   TextField "Screen title" at 783,728 size 496x50; Text 'Screen title'
   Bar "Bar_1" at 262,206 size 122x241; MinimumValue 0; MaximumValue 100
      ProcessValue <- "20_TANKS_IP_DATA_RIO_06_FIRST_TANK_BWT_LEVEL"
   Button "Button_48" at 273,396 size 100x25; TextOff 'DISABLED'
      on Release: function_efd93a16("Tank 6P Status", 168, 315, -1, 2, 1)
      Visibility <- "504_Tank Grouping_DB2020_GROUP of TANK 12"
   Circle "Circle_3" at 340,212 size 14x14
      Appearance <- "20_TANKS_IP_DATA_RIO_06_FIRST_TANK_BWT_LEVEL_HIHI"
   TextField "Text field_125" at 295,212 size 51x14; Text 'LS425-6P'
   Polyline "Polyline_1" at 261,205 size 123x240
      Visibility <- "504_Tank Grouping_DB2020_RUN TANK 12"
   TextField "Text field_64" at 288,273 size 74x20; Text 'Tank - 6P'
   Bar "Bar_2" at 394,206 size 122x241; MinimumValue 0; MaximumValue 100
      ProcessValue <- "20_TANKS_IP_DATA_RIO_05_FIRST_TANK_BWT_LEVEL"
   Button "Button_44" at 406,396 size 100x25; TextOff 'DISABLED'
      on Release: function_efd93a16("Tank 5P Status", 168, 315, -1, 2, 1)
      Visibility <- "504_Tank Grouping_DB2020_GROUP of TANK 10"
   Circle "Circle_4" at 472,212 size 14x14
      Appearance <- "20_TANKS_IP_DATA_RIO_05_FIRST_TANK_BWT_LEVEL_HIHI"
   TextField "Text field_124" at 427,212 size 51x14; Text 'LS425-5P'
   Polyline "Polyline_2" at 392,205 size 123x240
      Visibility <- "504_Tank Grouping_DB2020_RUN TANK 10"
   TextField "Text field_8" at 418,275 size 74x20; Text 'Tank - 5P'
   Bar "Bar_3" at 525,206 size 122x241; MinimumValue 0; MaximumValue 100
      ProcessValue <- "20_TANKS_IP_DATA_RIO_04_FIRST_TANK_BWT_LEVEL"
   Button "Button_40" at 537,395 size 100x25; TextOff 'DISABLED'
      on Release: function_efd93a16("Tank 4P Status", 168, 315, -1, 2, 1)
      Visibility <- "504_Tank Grouping_DB2020_GROUP of TANK 8"
   Circle "Circle_5" at 604,212 size 14x14
      Appearance <- "20_TANKS_IP_DATA_RIO_04_FIRST_TANK_BWT_LEVEL_HIHI"
   TextField "Text field_123" at 559,212 size 51x14; Text 'LS425-4P'
   Polyline "Polyline_3" at 525,205 size 123x240
      Visibility <- "504_Tank Grouping_DB2020_RUN TANK 8"
   TextField "Text field_9" at 553,275 size 74x20; Text 'Tank - 4P'
   Bar "Bar_4" at 657,206 size 122x241; MinimumValue 0; MaximumValue 100
      ProcessValue <- "20_TANKS_IP_DATA_RIO_03_FIRST_TANK_BWT_LEVEL"
   Button "Button_36" at 668,395 size 100x25; TextOff 'DISABLED'
      on Release: function_efd93a16("Tank 3P Status", 168, 315, -1, 0, 1)
      Visibility <- "504_Tank Grouping_DB2020_GROUP of TANK 6"
   Circle "Circle_7" at 736,212 size 14x14
      Appearance <- "20_TANKS_IP_DATA_RIO_03_FIRST_TANK_BWT_LEVEL_HIHI"
   TextField "Text field_122" at 691,212 size 51x14; Text 'LS425-3P'
   Polyline "Polyline_4" at 656,205 size 123x240
      Visibility <- "504_Tank Grouping_DB2020_RUN TANK 6"
   TextField "Text field_14" at 680,275 size 74x20; Text 'Tank - 3P'
   Bar "Bar_5" at 789,206 size 122x241; MinimumValue 0; MaximumValue 100
      ProcessValue <- "20_TANKS_IP_DATA_RIO_02_FIRST_TANK_BWT_LEVEL"
   Button "Button_32" at 802,396 size 100x25; TextOff 'DISABLED'
      on Release: function_efd93a16("Tank 2P Status", 168, 315, -1, 0, 1)
      Visibility <- "504_Tank Grouping_DB2020_GROUP of TANK 4"
   Circle "Circle_15" at 868,212 size 14x14
      Appearance <- "20_TANKS_IP_DATA_RIO_02_FIRST_TANK_BWT_LEVEL_HIHI"
   TextField "Text field_121" at 823,212 size 51x14; Text 'LS425-2P'
   Polyline "Polyline_5" at 789,205 size 123x240
      Visibility <- "504_Tank Grouping_DB2020_RUN TANK 4"
   TextField "Text field_15" at 816,275 size 74x20; Text 'Tank - 2P'
   Bar "Bar_6" at 922,205 size 122x241; MinimumValue 0; MaximumValue 100
      ProcessValue <- "20_TANKS_IP_DATA_RIO_01_SECOND_TANK_BWT_LEVEL"
   Button "Button_52" at 934,395 size 100x25; TextOff 'DISABLED'
      on Release: function_efd93a16("Tank 1P Status", 168, 315, -1, 0, 1)
      Visibility <- "504_Tank Grouping_DB2020_GROUP of TANK 2"
   Circle "Circle_16" at 999,211 size 14x14
      Appearance <- "20_TANKS_IP_DATA_RIO_01_SECOND_TANK_BWT_LEVEL_HIHI"
   TextField "Text field_120" at 955,211 size 51x14; Text 'LS425-1P'
   Polyline "Polyline_6" at 921,205 size 123x240
      Visibility <- "504_Tank Grouping_DB2020_RUN TANK 2"
   GraphicView "Graphic view_6" at 127,446 size 591x12; Picture "Graphic_151"
   TextField "Text field_16" at 947,275 size 74x20; Text 'Tank - 1P'
   Bar "Bar_7" at 1096,334 size 122x241; MinimumValue 0; MaximumValue 100
      ProcessValue <- "20_TANKS_IP_DATA_RIO_01_FIRST_TANK_BWT_LEVEL"
   Circle "Circle_24" at 1168,339 size 14x14
      Appearance <- "20_TANKS_IP_DATA_RIO_01_FIRST_TANK_BWT_LEVEL_HIHI"
   TextField "Text field_133" at 1139,339 size 35x14; Text 'LS425'
   Polyline "Polyline_14" at 1095,332 size 125x242
      Visibility <- "504_Tank Grouping_DB2020_RUN TANK 1"
   Button "Button_56" at 1110,524 size 100x25; TextOff 'DISABLED'
      on Release: function_efd93a16("Tank FP Status", 168, 315, -1, 0, 1)
      Visibility <- "504_Tank Grouping_DB2020_GROUP of TANK 1"
   TextField "Text field_17" at 1111,400 size 111x20; Text 'Fore PeakTank'
   Bar "Bar_8" at 922,458 size 122x258; MinimumValue 0; MaximumValue 100
      ProcessValue <- "20_TANKS_IP_DATA_RIO_01_THIRD_TANK_BWT_LEVEL"
   Button "Button_54" at 933,661 size 100x25; TextOff 'DISABLED'
      on Release: function_efd93a16("Tank 1S Status", 168, 315, -1, 0, 1)
      Visibility <- "504_Tank Grouping_DB2020_GROUP of TANK 3"
   Circle "Circle_23" at 1000,464 size 14x14
      Appearance <- "20_TANKS_IP_DATA_RIO_01_THIRD_TANK_BWT_LEVEL_HIHI"
   TextField "Text field_126" at 955,465 size 51x14; Text 'LS422-1S'
   Polyline "Polyline_7" at 921,458 size 123x259
      Visibility <- "504_Tank Grouping_DB2020_RUN TANK 3"
   TextField "Text field_10" at 950,618 size 74x20; Text 'Tank - 1S'
   Bar "Bar_9" at 790,459 size 122x258; MinimumValue 0; MaximumValue 100
      ProcessValue <- "20_TANKS_IP_DATA_RIO_02_SECOND_TANK_BWT_LEVEL"
   Button "Button_34" at 801,662 size 100x25; TextOff 'DISABLED'
      on Release: function_efd93a16("Tank 2S Status", 168, 315, -1, 0, 1)
      Visibility <- "504_Tank Grouping_DB2020_GROUP of TANK 5"
   Circle "Circle_22" at 868,465 size 14x14
      Appearance <- "20_TANKS_IP_DATA_RIO_02_SECOND_TANK_BWT_LEVEL_HIHI"
   TextField "Text field_127" at 823,466 size 51x14; Text 'LS422-2S'
   Polyline "Polyline_8" at 789,458 size 123x259
      Visibility <- "504_Tank Grouping_DB2020_RUN TANK 5"
   TextField "Text field_11" at 817,618 size 74x20; Text 'Tank - 2S'
   Bar "Bar_10" at 659,460 size 122x258; MinimumValue 0; MaximumValue 100
      ProcessValue <- "20_TANKS_IP_DATA_RIO_03_SECOND_TANK_BWT_LEVEL"
   Button "Button_38" at 669,663 size 100x25; TextOff 'DISABLED'
      on Release: function_efd93a16("Tank 3S Status", 168, 315, -1, 0, 1)
      Visibility <- "504_Tank Grouping_DB2020_GROUP of TANK 7"
   Circle "Circle_21" at 736,467 size 14x14
      Appearance <- "20_TANKS_IP_DATA_RIO_03_SECOND_TANK_BWT_LEVEL_HIHI"
   TextField "Text field_128" at 691,468 size 51x14; Text 'LS422-3S'
   Polyline "Polyline_9" at 658,458 size 123x259
      Visibility <- "504_Tank Grouping_DB2020_RUN TANK 7"
   TextField "Text field_12" at 690,618 size 74x20; Text 'Tank - 3S'
   Bar "Bar_11" at 526,459 size 122x258; MinimumValue 0; MaximumValue 100
      ProcessValue <- "20_TANKS_IP_DATA_RIO_04_SECOND_TANK_BWT_LEVEL"
   Button "Button_42" at 537,662 size 100x25; TextOff 'DISABLED'
      on Release: function_efd93a16("Tank 4S Status", 168, 315, -1, 2, 1)
      Visibility <- "504_Tank Grouping_DB2020_GROUP of TANK 9"
   Circle "Circle_19" at 604,466 size 14x14
      Appearance <- "20_TANKS_IP_DATA_RIO_04_SECOND_TANK_BWT_LEVEL_HIHI"
   TextField "Text field_129" at 559,467 size 51x14; Text 'LS422-4S'
   Polyline "Polyline_10" at 525,458 size 123x259
      Visibility <- "504_Tank Grouping_DB2020_RUN TANK 9"
   TextField "Text field_13" at 554,618 size 74x20; Text 'Tank - 4S'
   Bar "Bar_12" at 394,459 size 122x258; MinimumValue 0; MaximumValue 100
      ProcessValue <- "20_TANKS_IP_DATA_RIO_05_SECOND_TANK_BWT_LEVEL"
   Button "Button_46" at 405,662 size 100x25; TextOff 'DISABLED'
      on Release: function_efd93a16("Tank 5S Status", 168, 315, -1, 2, 1)
      Visibility <- "504_Tank Grouping_DB2020_GROUP of TANK 11"
   Circle "Circle_18" at 472,465 size 14x14
      Appearance <- "20_TANKS_IP_DATA_RIO_05_SECOND_TANK_BWT_LEVEL_HIHI"
   TextField "Text field_130" at 427,466 size 51x14; Text 'LS422-5S'
   Polyline "Polyline_11" at 393,458 size 123x259
      Visibility <- "504_Tank Grouping_DB2020_RUN TANK 11"
   TextField "Text field_18" at 424,618 size 74x20; Text 'Tank - 5S'
   Bar "Bar_13" at 262,460 size 122x258; MinimumValue 0; MaximumValue 100
      ProcessValue <- "20_TANKS_IP_DATA_RIO_06_SECOND_TANK_BWT_LEVEL"
   Button "Button_50" at 273,663 size 100x25; TextOff 'DISABLED'
      on Release: function_efd93a16("Tank 6S Status", 168, 315, -1, 2, 1)
      Visibility <- "504_Tank Grouping_DB2020_GROUP of TANK 13"
   Circle "Circle_17" at 340,467 size 14x14
      Appearance <- "20_TANKS_IP_DATA_RIO_06_SECOND_TANK_BWT_LEVEL_HIHI"
   TextField "Text field_131" at 295,468 size 51x14; Text 'LS422-6S'
   Polyline "Polyline_12" at 261,458 size 123x258
      Visibility <- "504_Tank Grouping_DB2020_RUN TANK 13"
   TextField "Text field_19" at 290,618 size 74x20; Text 'Tank - 6S'
   Bar "Bar_14" at 39,324 size 119x258; Unit %; MinimumValue 0; MaximumValue 100
      ProcessValue <- "20_TANKS_IP_DATA_RIO_07_FIRST_TANK_BWT_LEVEL"
   Circle "Circle_25" at 108,330 size 14x14
      Appearance <- "20_TANKS_IP_DATA_RIO_07_FIRST_TANK_BWT_LEVEL_HIHI"
   TextField "Text field_132" at 79,330 size 35x14; Text 'LS425'
   Polyline "Polyline_13" at 38,324 size 121x259
      Visibility <- "504_Tank Grouping_DB2020_RUN TANK 14"
   Button "Button_58" at 48,527 size 100x25; TextOff 'DISABLED'
      on Release: function_efd93a16("Tank AP Status", 168, 315, -1, 2, 1)
      Visibility <- "504_Tank Grouping_DB2020_GROUP of TANK 14"
   Button "HmiScreenItemData_6" at 1043,144 size 116x50; TextOn 'Back'; TextOff 'Tank Status'
      on Release: ActivateScreen("Balast Water Treatment Plant", 0)
   Button "Button_2" at 252,437 size 37x30; TextOff 'DB&B'
      on Release: function_efd93a16("Double Block & Bleed Valve Monitoring", 250, 250, -1, -1, 1)
      Appearance <- "10_DI_DATA_CV407_OPN"
   TextField "Text field_65" at 190,398 size 46x25; Text 'PGC'
   TextField "Text field_75" at 183,480 size 60x20; Text 'Disabled'
   TextField "Text field_76" at 183,480 size 60x20; Text 'Enabled'
      Visibility <- "10_DI_DATA_E_400_RUN"
   GraphicView "Graphic view_76" at 185,421 size 57x55; Picture "Graphic_251"
   Button "Button_6" at 179,402 size 70x105; TextOff 'Text'
      on Release: ActivateScreen("PGC System", 0)
   TextField "Text field_20" at 53,396 size 103x20; Text 'Aft PeakTank'
   GraphicView "Graphic view_108" at 4,683 size 96x48; Picture "Left Arow"
   Button "HmiScreenItemData_14" at 3,660 size 106x93; TextOn 'Back'; TextOff 'Text'
      on Press: ActivateScreen("Inert Gas Conditioning Plant", 0)
   IOField "I/O field_1" at 68,460 size 84x25; FormatPattern 99.99; Unit m
      ProcessValue <- "Data_From_WBT_Level_APT m"
   IOField "I/O field_2" at 285,331 size 84x25; FormatPattern 99.99; Unit m
      ProcessValue <- "Data_From_WBT_Level_WBT_6P m"
   IOField "I/O field_3" at 418,331 size 84x25; FormatPattern 99.99; Unit m
      ProcessValue <- "Data_From_WBT_Level_WBT_5P m"
   IOField "I/O field_4" at 550,331 size 84x25; FormatPattern 99.99; Unit m
      ProcessValue <- "Data_From_WBT_Level_WBT_4P m"
   IOField "I/O field_5" at 681,331 size 84x25; FormatPattern 99.99; Unit m
      ProcessValue <- "Data_From_WBT_Level_WBT_3P m"
   IOField "I/O field_6" at 815,331 size 84x25; FormatPattern 99.99; Unit m
      ProcessValue <- "Data_From_WBT_Level_WBT_2P m"
   IOField "I/O field_7" at 949,331 size 84x25; FormatPattern 99.99; Unit m
      ProcessValue <- "Data_From_WBT_Level_WBT_1P m"
   IOField "I/O field_8" at 1124,459 size 84x25; FormatPattern 99.99; Unit m
      ProcessValue <- "Data_From_WBT_Level_FPT m"
   IOField "I/O field_9" at 945,555 size 84x25; FormatPattern 99.99; Unit m
      ProcessValue <- "Data_From_WBT_Level_WBT_1S m"
   IOField "I/O field_10" at 816,556 size 84x25; FormatPattern 99.99; Unit m
      ProcessValue <- "Data_From_WBT_Level_WBT_2S m"
   IOField "I/O field_11" at 685,558 size 84x25; FormatPattern 99.99; Unit m
      ProcessValue <- "Data_From_WBT_Level_WBT_3S m"
   IOField "I/O field_12" at 553,557 size 84x25; FormatPattern 99.99; Unit m
      ProcessValue <- "Data_From_WBT_Level_WBT_4S m"
   IOField "I/O field_13" at 418,558 size 84x25; FormatPattern 99.99; Unit m
      ProcessValue <- "Data_From_WBT_Level_WBT_5S m"
   IOField "I/O field_14" at 287,559 size 84x25; FormatPattern 99.99; Unit m
      ProcessValue <- "Data_From_WBT_Level_WBT_6S m"
   Button "Button_88" at 34,324 size 127x264; TextOff 'Text'
      on Release: function_efd93a16("Tank AP Status", 168, 315, -1, 0, 1)
      Appearance <- "504_Tank Grouping_DB2020_RUN TANK 14"
   Button "Button_86" at 259,458 size 126x260; TextOff 'Text'
      on Release: function_efd93a16("Tank 6S Status", 168, 315, -1, 0, 1)
      Appearance <- "504_Tank Grouping_DB2020_RUN TANK 13"
   Button "Button_79" at 391,457 size 126x262; TextOff 'Text'
      on Release: function_efd93a16("Tank 5S Status", 168, 315, -1, 0, 1)
      Appearance <- "504_Tank Grouping_DB2020_RUN TANK 11"
   Button "Button_77" at 523,457 size 126x262; TextOff 'Text'
      on Release: function_efd93a16("Tank 4S Status", 168, 315, -1, 0, 1)
      Appearance <- "504_Tank Grouping_DB2020_RUN TANK 9"
   Button "Button_74" at 657,457 size 126x262; TextOff 'Text'
      on Release: function_efd93a16("Tank 3S Status", 168, 315, -1, 0, 1)
      Appearance <- "504_Tank Grouping_DB2020_RUN TANK 7"
   Button "Button_70" at 788,457 size 126x262; TextOff 'Text'
      on Release: function_efd93a16("Tank 2S Status", 168, 315, -1, 0, 1)
      Appearance <- "504_Tank Grouping_DB2020_RUN TANK 5"
   Button "Button_66" at 921,457 size 126x261; TextOff 'Text'
      on Release: function_efd93a16("Tank 1S Status", 168, 315, -1, 0, 1)
      Appearance <- "504_Tank Grouping_DB2020_RUN TANK 3"
   Button "Button_61" at 1093,328 size 130x248; TextOff 'Text'
      on Release: function_efd93a16("Tank FP Status", 168, 315, -1, 0, 1)
      Appearance <- "504_Tank Grouping_DB2020_RUN TANK 1"
   Button "Button_62" at 919,205 size 126x242; TextOff 'Text'
      on Release: function_efd93a16("Tank 1P Status", 168, 315, -1, 0, 1)
      Appearance <- "504_Tank Grouping_DB2020_RUN TANK 2"
   Button "Button_68" at 789,202 size 126x246; TextOff 'Text'
      on Release: function_efd93a16("Tank 2P Status", 168, 315, -1, 0, 1)
      Appearance <- "504_Tank Grouping_DB2020_RUN TANK 4"
   Button "Button_72" at 654,205 size 126x242; TextOff 'Text'
      on Release: function_efd93a16("Tank 3P Status", 168, 315, -1, 0, 1)
      Appearance <- "504_Tank Grouping_DB2020_RUN TANK 6"
   Button "Button_76" at 524,205 size 126x243; TextOff 'Text'
      on Release: function_efd93a16("Tank 4P Status", 168, 315, -1, 0, 1)
      Appearance <- "504_Tank Grouping_DB2020_RUN TANK 8"
   Button "Button_78" at 392,206 size 126x241; TextOff 'Text'
      on Release: function_efd93a16("Tank 5P Status", 168, 315, -1, 0, 1)
      Appearance <- "504_Tank Grouping_DB2020_RUN TANK 10"
   Button "Button_84" at 259,204 size 126x244; TextOff 'Text'
      on Release: function_efd93a16("Tank 6P Status", 168, 315, -1, 0, 1)
      Appearance <- "504_Tank Grouping_DB2020_RUN TANK 12"
   Group "Group_5" at 664,46 size 45x27; FormatPattern 999
   Group "Group_1" at 711,46 size 50x27; FormatPattern 999; Unit h
   Group "Group_2" at 605,46 size 57x27; FormatPattern 999; Unit h
   Button "HmiScreenItemData_5" at 180,144 size 116x50; TextOn 'Back'; TextOff 'Tank Status'
      on Release: function_efd93a16("Tank Status", 400, 250, -1, -1, 1)
   Button "Button_10" at 14,93 size 153x55; TextOff 'Text'
      on Release: function_efd93a16("Salinity - Acceptance", 168, 315, -1, 0, 1)
      Visibility <- "2068_Sys_Status_Data_SAL_VALID"
   Button "Button_12" at 14,93 size 153x53; TextOff 'Text'
      on Release: function_efd93a16("Tank Times", 300, 200, -1, 0, 1)
      Visibility <- "2068_Sys_Status_Data_Times Visibil"
   Button "Button_59" at 298,44 size 240x30; TextOn 'TB3 Enabled'; TextOff 'BWT System Shutting Down'
      Visibility <- "2110_BTCS_CNTRL_DB_BTCS_STATE"
   Button "Button_60" at 299,44 size 240x30; TextOn 'TB3 Enabled'; TextOff 'BWT System Enabled'
      Visibility <- "2110_BTCS_CNTRL_DB_BTCS_STATE"
   IOField "I/O field_29" at 664,46 size 45x27; FormatPattern 99; Unit h
      ProcessValue <- "Sequence Times_DB_Treatment Timer_Hours Left"
      Visibility <- "2110_BTCS_CNTRL_DB_BTCS_STATE"
   IOField "I/O field_30" at 664,46 size 45x27; FormatPattern 99; Unit h
      ProcessValue <- "Sequence Times_DB_Pre-Dwell Timer_Hours Left"
      Visibility <- "2110_BTCS_CNTRL_DB_BTCS_STATE"
   IOField "I/O field_15" at 711,46 size 50x27; FormatPattern 99; Unit m
      ProcessValue <- "Sequence Times_DB_Treatment Timer_Minutes Left"
      Visibility <- "2110_BTCS_CNTRL_DB_BTCS_STATE"
   IOField "I/O field_16" at 711,46 size 50x27; FormatPattern 99; Unit m
      ProcessValue <- "Sequence Times_DB_Pre-Dwell Timer_Minutes Left"
      Visibility <- "2110_BTCS_CNTRL_DB_BTCS_STATE"
   IOField "I/O field_17" at 605,46 size 57x27; FormatPattern 999; Unit d
      ProcessValue <- "Sequence Times_DB_Treatment Timer_Days Left"
      Visibility <- "2110_BTCS_CNTRL_DB_BTCS_STATE"
   IOField "I/O field_18" at 605,46 size 57x27; FormatPattern 999; Unit d
      ProcessValue <- "Sequence Times_DB_Pre-Dwell Timer_Days Left"
      Visibility <- "2110_BTCS_CNTRL_DB_BTCS_STATE"

screen "PGC System" 1280x800, template "Template"
   Button "HmiScreenItemData_1" at -189,1 size 150x43; TextOn 'Back'; TextOff 'Main Index'
      on Release: ActivateScreen("02 Main Index", 0)
   Gauge "Gauge_1" at 454,351 size 184x184; CaptionText 'Pressure'; UnitText 'Bar'
      ProcessValue <- "12_AI_Data_E_400_PT002_SCALED"
      MaximumValue <- "84_Setpoints_E400_PT002_HighHigh"
   TextField "Text field_20" at 187,312 size 324x26; Text 'Process Gas Discharge Pressure'
   TextField "Text field_7" at 221,72 size 326x26; Text 'Process Gas Compressor Control'
   TextField "Text field_10" at 119,405 size 243x20; Text 'Process Gas Discharge Pressure'
   TextField "Text field_17" at 119,464 size 217x20; Text 'Discharge Pressure Setpoint'
   Button "Button_8" at 117,115 size 240x30; TextOn 'TB3 Enabled'; TextOff 'PGC System Not Running OK'
      Visibility <- "10_DI_DATA_E_400_RUN"
   Button "HmiScreenItemData_12" at 141,237 size 69x51; TextOn 'Back'; TextOff 'Reset'; Authorization "Operate"
      on Press: function_b14e0dd5("140_PGC_HRS_RUN_DB_RST", 0)
   IOField "I/O field_10" at 70,236 size 66x25; FormatPattern 9999; Unit  h
      ProcessValue <- "140_PGC_HRS_RUN_DB_SRV_HRS"
   TextField "Text field_22" at 36,238 size 37x20; Text 'Run'
   TextField "Text field_23" at 36,268 size 37x20; Text 'Set'
   TextField "Text field_24" at 79,212 size 100x20; Text 'Service Hour'
   IOField "I/O field_13" at 222,249 size 75x25; FormatPattern 99999; Unit h
      ProcessValue <- "140_PGC_HRS_RUN_DB_HRS"
   IOField "I/O field_14" at 299,249 size 40x25; FormatPattern 99; Unit m
      ProcessValue <- "140_PGC_HRS_RUN_DB_MINS"
   IOField "I/O field_15" at 341,249 size 40x25; FormatPattern 99; Unit s
      ProcessValue <- "140_PGC_HRS_RUN_DB_SECS"
   Button "Button_7" at 654,76 size 57x25; TextOn 'Alarm'; TextOff 'Service'
      Visibility <- "140_PGC_HRS_RUN_DB_SRVC"
      Appearance <- "140_PGC_HRS_RUN_DB_SRVC"
   Button "Button_15" at 187,173 size 57x25; TextOn 'Enabled'; TextOff 'Disabled'
   Button "Button_16" at 341,173 size 64x25; TextOn 'Alarm'; TextOff 'Text'
   TextField "Text field_14" at 44,175 size 115x20; Text 'PG Compressor'
   TextField "Text field_15" at 191,151 size 60x18; Text 'Enabled'
   TextField "Text field_16" at 266,151 size 64x18; Text 'Running'
   TextField "Text field_18" at 343,150 size 78x18; Text 'Shutdown'
   Button "Button_1" at 264,173 size 57x25; TextOn 'Enabled'; TextOff 'Stopped'
   TextField "Text field_32" at 187,173 size 57x25; Text 'Enabled'
      Visibility <- "10_DI_DATA_E_400_SHTDN"
   TextField "Text field_2" at 264,173 size 57x25; Text 'Running'
      Visibility <- "10_DI_DATA_E_400_RUN"
   Button "Button_3" at 341,173 size 64x25; TextOn 'Enabled'; TextOff 'Normal'
   Button "Button_2" at 341,173 size 69x25; TextOn 'Alarm'; TextOff 'Shutdown'
      Visibility <- "10_DI_DATA_E_400_NOK"
      Appearance <- "10_DI_DATA_E_400_NOK"
   Gauge "Gauge_2" at 454,588 size 184x184; UnitText '°C'; CaptionText 'Temperature'
      ProcessValue <- "12_AI_Data_E_400_TE002_SCALED"
      MaximumValue <- "84_Setpoints_E400_TT002_HighHigh"
   TextField "Text field_1" at 187,549 size 365x26; Text 'Process Gas Discharge Temperature'
   TextField "Text field_3" at 119,641 size 178x20; Text 'Discharge Temperature'
   TextField "Text field_4" at 109,699 size 246x20; Text 'Discharge Temperature Setpoint'
   IOField "I/O field_2" at 332,403 size 66x25; FormatPattern 9.99; Unit  Bar
      ProcessValue <- "12_AI_Data_E_400_PT002_SCALED"
   IOField "I/O field_1" at 334,638 size 66x25; FormatPattern 999; Unit  °C
      ProcessValue <- "12_AI_Data_E_400_TE002_SCALED"
   Button "HmiScreenItemData_11" at 3,1 size 150x43; TextOn 'IGG Plant'; TextOff 'GCU Plant'
      on Release: ActivateScreen("Inert Gas Conditioning Plant", 0)
   IOField "I/O field_3" at 332,462 size 66x25; Authorization "Commissioning"; FormatPattern 9.99; Unit  Bar
      ProcessValue <- "84_Setpoints_E400_PT002_HighHigh"
   IOField "I/O field_4" at 334,697 size 66x25; Authorization "Commissioning"; FormatPattern 999; Unit  °C
      ProcessValue <- "84_Setpoints_E400_TT002_HighHigh"
   GraphicView "Graphic view_1" at 514,109 size 192x199; Picture "Graphic_251"
   Button "HmiScreenItemData_3" at 1125,1 size 150x43; TextOn 'I&A Compressor Ok'; TextOff 'Back'
      on Release: function_efd93a16()
   TextField "Text field_5" at 222,226 size 160x25; Text 'Total Run Time'
   TextField "Text field_6" at 818,74 size 312x26; Text 'Process Gas Compressor Purge'
   TextField "Text field_8" at 717,177 size 263x20; Text 'Process Gas Compresor Stop Delay'
   TextField "Text field_11" at 716,111 size 305x20; Text 'Combustion Air Blower after Start Delay'
   IOField "I/O field_7" at 993,109 size 66x25; FormatPattern 999; Unit s
      ProcessValue <- "PGC Flush_DB_CAB after Start Delay"
   TextField "Text field_12" at 716,144 size 208x20; Text 'Combustion Air Blower RPM'
   IOField "I/O field_8" at 993,142 size 66x25; FormatPattern 999; Unit RPM
      ProcessValue <- "PGC Flush_DB_CAB RPM Cmnd"
   Button "HmiScreenItemData_2" at 982,285 size 82x35; TextOn 'Back'; TextOff 'Override'; Authorization "Operating Mode"
      on Press: function_b14e0dd5("PGC Flush_DB_Override", 0)
      Appearance <- "PGC Flush_DB_Flip Flop_Override_Output"
   TextField "Text field_9" at 1068,149 size 91x21; Text 'Running'
      Appearance <- "PGC Flush_DB_Running"
   TextField "Text field_13" at 1068,129 size 91x21; Text 'Enabled'
      Appearance <- "PGC Flush_DB_Activate"
   TextField "Text field_19" at 1068,329 size 91x21; Text 'Done'
      Appearance <- "PGC Flush_DB_Done"
   TextField "Text field_21" at 1068,169 size 91x21; Text 'Open CV405'
      Appearance <- "PGC Flush_DB_CV405 Open"
   TextField "Text field_25" at 1068,189 size 91x21; Text 'Open CV401'
      Appearance <- "PGC Flush_DB_CV401 Open"
   TextField "Text field_26" at 1068,209 size 91x21; Text 'Open CV431'
      Appearance <- "PGC Flush_DB_CV431 Open"
   TextField "Text field_27" at 1068,249 size 91x21; Text 'Close CV441'
      Appearance <- "PGC Flush_DB_CV431 Open"
   TextField "Text field_28" at 1068,269 size 91x21; Text 'Start CAB'
      Appearance <- "PGC Flush_DB_CAB Start"
   TextField "Text field_29" at 1068,289 size 91x21; Text 'Mdlt CV403'
      Appearance <- "PGC Flush_DB_CV403 Modulate"
   TextField "Text field_30" at 1068,309 size 91x21; Text 'Stop PGC'
      Appearance <- "PGC Flush_DB_Stop PGC"
   IOField "I/O field_37" at 890,604 size 90x29; Authorization "Commissioning"; FormatPattern 999; Unit  step
      ProcessValue <- "2110_BTCS_CNTRL_DB_BTCS_STEP"
   Button "HmiScreenItemData_10" at 749,604 size 137x29; TextOn 'Back'; TextOff 'BWTS Step'
   Button "HmiScreenItemData_51" at 749,671 size 137x29; TextOn 'Back'; TextOff 'BWTS State'
   Button "HmiScreenItemData_54" at 749,633 size 495x29; TextOn 'Back'; TextOff 'IGG STEP'; TextList "STEP LIST BTCS"
      ProcessValue <- "2110_BTCS_CNTRL_DB_BTCS_STEP"
   Button "HmiScreenItemData_55" at 749,700 size 495x29; TextOn 'Back'; TextOff 'IGG STEP'; TextList "STATE LIST BTCS"
      ProcessValue <- "2110_BTCS_CNTRL_DB_BTCS_STATE"
   IOField "I/O field_38" at 890,671 size 90x29; Authorization "Commissioning"; FormatPattern 9; Unit  state
      ProcessValue <- "2110_BTCS_CNTRL_DB_BTCS_STATE"
   TextField "Text field_31" at 716,210 size 149x20; Text 'PGC Purge Duration'
   IOField "I/O field_6" at 993,208 size 66x25; FormatPattern 999; Unit m
      ProcessValue <- "PGC Flush_DB_PGC Purge Duration"
   TextField "Text field_33" at 1068,229 size 91x21; Text 'Open CV403'
      Appearance <- "PGC Flush_DB_CV403 Open"
   TextField "Text field_34" at 768,296 size 175x18; Text 'Purge Request Simulate'
      Visibility <- "user_group"
   Switch "Switch_1" at 726,288 size 32x29; CaptionText 'Switch'; TextOn 'ON'; TextOff 'OFF'; Authorization "User administration"; PictureOff "Design_5_PilotLight_Green_Off"; PictureOn "Design_5_PilotLight_Green_On"
      on Change: InvertBit("Sequence Times_DB_Treatment Timer_Enable")
      Visibility <- "user_group"
      ProcessValue <- "19_AUTO_CMNDS_Data_Purge Rqst Simulate"
   TextField "Text field_35" at 1160,149 size 106x21; Text 'Running'
      Appearance <- "PGC Flush_DB_Running"
   TextField "Text field_36" at 1160,129 size 106x21; Text 'Enabled'
      Appearance <- "PGC Flush_DB_Activate"
   TextField "Text field_37" at 1160,329 size 106x21; Text 'Done'
      Appearance <- "100_GCU_AUTO_SEQ_DB_CRNT_STEP"
   TextField "Text field_38" at 1160,169 size 106x21; Text 'Opened CV405'
      Appearance <- "1405_PID_CV405_ManualEnable"
   TextField "Text field_39" at 1160,189 size 106x21; Text 'Opened CV401'
      Appearance <- "PGC Flush_DB_CV401 Opened"
   TextField "Text field_40" at 1160,209 size 106x21; Text 'Opened CV431'
      Appearance <- "PGC Flush_DB_CV431 Opened"
   TextField "Text field_41" at 1160,249 size 106x21; Text 'Closed CV441'
      Appearance <- "PGC Flush_DB_CV441 Closed"
   TextField "Text field_42" at 1160,269 size 106x21; Text 'Started CAB'
      Appearance <- "PGC Flush_DB_CAB Started"
   TextField "Text field_43" at 1160,289 size 106x21; Text 'Mdling CV403'
      Appearance <- "1403_PID_300CV403_ModeActivate"
   TextField "Text field_44" at 1160,309 size 106x21; Text 'Stoped PGC'
      Appearance <- "PGC Flush_DB_PGC Stoped"
   TextField "Text field_45" at 1160,229 size 106x21; Text 'Opened CV403'
      Appearance <- "1403_PID_300CV403_ManualEnable"
   TextField "Text field_46" at 711,332 size 173x20; Text 'Air / Inert Gas Pressure'
   Button "Button_9" at 1001,329 size 57x25; TextOn 'Enabled'; TextOff 'Text'
   TextField "Text field_47" at 710,366 size 277x20; Text 'Air / Inert Gas Pressure Setpoint (Pre-Ignition)'
   Button "Button_11" at 1001,364 size 57x25; TextOn 'Enabled'; TextOff 'Text'
   TextField "Text field_48" at 718,498 size 182x20; Text 'Modulating Valve Position'
   TextField "Text field_49" at 709,399 size 278x20; Text 'Air / Inert Gas Pressure Setpoint (Main-Ignition)'
   Button "Button_10" at 1001,397 size 57x25; TextOn 'Enabled'; TextOff 'Text'
   IOField "I/O field_9" at 993,329 size 66x25; FormatPattern 999; Unit  mbar
      ProcessValue <- "12_AI_Data_PIT402_SCALED"
   IOField "I/O field_12" at 993,364 size 66x25; Authorization "Commissioning"; FormatPattern 999; Unit  mbar
      ProcessValue <- "84_Setpoints_PIT402_Pilot_Target"
   IOField "I/O field_16" at 993,495 size 66x25; FormatPattern 999; Unit  %
      ProcessValue <- "16_AQ_Data_CV403_CNTRL"
   IOField "I/O field_17" at 993,462 size 66x25; FormatPattern 999; Unit  mBar
      ProcessValue <- "19_AUTO_CMNDS_Data_PIT402_Target"
      Appearance <- "19_AUTO_CMNDS_Data_PIT402_Target"
   IOField "I/O field_18" at 993,396 size 66x25; Authorization "Commissioning"; FormatPattern 999; Unit  mbar
      ProcessValue <- "84_Setpoints_PIT402_Main_Target"
   TextField "Text field_50" at 1068,497 size 58x20; Text 'Opened'
   TextField "Text field_51" at 711,465 size 266x20; Text 'Air / Inert Gas Pressure Setpoint (Current)'
   TextField "Text field_52" at 709,432 size 278x20; Text 'Air / Inert Gas Pressure Setpoint (Post-Ignition)'
   Button "Button_4" at 1001,430 size 57x25; TextOn 'Enabled'; TextOff 'Text'
   IOField "I/O field_19" at 993,429 size 66x25; Authorization "Commissioning"; FormatPattern 999; Unit  mbar
      ProcessValue <- "84_Setpoints_PIT401_Post_Target_Max"
   TextField "Text field_53" at 1079,107 size 73x20; Text 'Command'
   TextField "Text field_54" at 1182,107 size 73x20; Text 'Feedback'
   IOField "I/O field_20" at 70,266 size 66x25; Authorization "Commissioning"; FormatPattern 9999; Unit h
      ProcessValue <- "140_PGC_HRS_RUN_DB_SHRS_IP"
   TextField "Text field_55" at 716,243 size 168x20; Text 'Temperature Setpoint'
   IOField "I/O field_11" at 993,241 size 66x25; FormatPattern 999; Unit  °C
      ProcessValue <- "PGC Flush_DB_Temperature Setpoint"
   Button "HmiScreenItemData_19" at 749,567 size 495x29; TextOn 'Back'; TextOff 'IGG STEP'; TextList "STEP LIST_GCU"
      ProcessValue <- "100_GCU_AUTO_SEQ_DB_CRNT_STEP"
   IOField "I/O field_21" at 890,537 size 90x29; Authorization "Commissioning"; FormatPattern 999; Unit  Step
      ProcessValue <- "100_GCU_AUTO_SEQ_DB_CRNT_STEP"
   Button "HmiScreenItemData_9" at 749,536 size 100x30; TextOn 'Back'; TextOff 'GCU PLC'
   Button "HmiScreenItemData_16" at 238,742 size 83x29; TextOn 'Back'; TextOff 'Temp-Trends'
      on Click: function_efd93a16("PGC Temperature Trends", 200, 100, -1, -1, 1)
   IOField "I/O field_22" at 993,175 size 66x25; FormatPattern 999; Unit m
      ProcessValue <- "PGC Flush_DB_PGC Stop Delay"

screen "Fresh Water System" 1280x800, template "Template"
   GraphicView "Graphic view_29" at 858,564 size 26x29; Picture "Graphic_155"
   Bar "Bar_1" at 145,436 size 311x274; Unit  %; MinimumValue 0; MaximumValue 100
      ProcessValue <- "12_AI_Data_LIT305_SCALED"
   GraphicView "Graphic view_15" at 640,691 size 216x15; Picture "Graphic_156"
   GraphicView "Graphic view_22" at 468,691 size 71x15; Picture "Graphic_156"
   TextField "Text field_1" at 262,720 size 73x32; Text 'IBC-2 Bulk Tank'
   GraphicView "Graphic view_3" at 454,688 size 6x20; Picture "Graphic_113"
   TextField "Text field_4" at 442,89 size 268x26; Text 'Fresh Water Pump Control'
   IOField "I/O field_2" at 646,242 size 65x25; FormatPattern 99999; Unit  h
      ProcessValue <- "P305_Functioning Hours_IDB_Hours Functioning Out"
   TextField "Text field_5" at 616,244 size 37x20; Text 'Run'
   TextField "Text field_6" at 616,275 size 37x20; Text 'Set'
   TextField "Text field_9" at 659,141 size 100x20; Text 'Service Hour'
   Button "HmiScreenItemData_10" at 639,169 size 178x34; TextOn 'Back'; TextOff 'Text'
   IOField "I/O field_4" at 689,173 size 40x25; FormatPattern 99; Unit h
      ProcessValue <- "82_To_HMI_P305 FW Pump Run Hours"
   IOField "I/O field_5" at 730,173 size 40x25; FormatPattern 99; Unit m
      ProcessValue <- "P305_Functioning Hours_IDB_Minutes"
   IOField "I/O field_6" at 771,173 size 40x25; FormatPattern 99; Unit s
      ProcessValue <- "P305_Functioning Hours_IDB_Seconds"
   Button "Button_4" at 776,90 size 57x25; TextOn 'Alarm'; TextOff 'Service'
      Visibility <- "P305_Functioning Hours_IDB_Service Time bit"
   Button "Button_9" at 374,166 size 57x25; TextOn 'Enabled'; TextOff 'Disabled'
   Button "Button_11" at 528,166 size 64x25; TextOn 'Alarm'; TextOff 'Text'
   TextField "Text field_10" at 231,168 size 140x20; Text 'Fresh Water Pump'
   TextField "Text field_8" at 378,144 size 60x18; Text 'Enabled'
   TextField "Text field_17" at 453,144 size 64x18; Text 'Running'
   TextField "Text field_20" at 533,144 size 58x18; Text 'Tripped'
      Visibility <- "10 DI_DATA_P305_TRIPPED(1)"
   Button "Button_12" at 451,166 size 57x25; TextOn 'Enabled'; TextOff 'Stopped'
   TextField "Text field_26" at 374,166 size 57x25; Text 'Enabled'
      Visibility <- "14_DQ_Data_P305ControlOut"
   TextField "Text field_27" at 448,166 size 64x25; Text 'Running'
      Visibility <- "10 DI_DATA_P305_ENBLD"
   GraphicView "Graphic view_12" at 396,411 size 20x26; Picture "Graphic_36"
   TextField "Text field_11" at 421,411 size 60x18; Text 'LIT-305'
   GraphicView "Graphic view_13" at 518,691 size 71x15; Picture "Graphic_156"
   GraphicView "Graphic view_11" at 456,691 size 15x15; Picture "Graphic_156"
   GraphicView "Graphic view_27" at 846,676 size 25x29; Picture "Graphic_153"
   GraphicView "Graphic view_28" at 858,581 size 13x101; Picture "Graphic_152"
   GraphicView "Graphic view_30" at 876,702 size 146x15; Picture "Graphic_156"
   GraphicView "Graphic view_31" at 870,564 size 152x15; Picture "Graphic_156"
   GraphicView "Graphic view_32" at 858,688 size 26x29; Picture "Graphic_166"
   TextField "Text field_15" at 550,746 size 133x32; Text 'P-305 Fresh Water Pump'
   Button "Button_1" at 528,166 size 64x25; TextOn 'Alarm'; TextOff 'Tripped'
      Visibility <- "10 DI_DATA_P305_TRIPPED"
      Appearance <- "10 DI_DATA_P305_TRIPPED"
   IOField "I/O field_13" at 376,388 size 63x18; FormatPattern 99.9; Unit  %
      ProcessValue <- "12_AI_Data_LIT305_SCALED"
   TextField "Text field_22" at 1059,560 size 168x21; Text 'Fresh Water Supply To GCU'
   TextField "Text field_3" at 1059,699 size 168x21; Text 'Fresh Water Supply To IGG'
   Button "HmiScreenItemData_9" at 721,243 size 69x51; TextOn 'Back'; TextOff 'SReset'; Authorization "Operating Mode"
      on Press: function_b14e0dd5("82_To_HMI_P305 FW Pump Reset Hours", 0)
   GraphicView "Graphic view_1" at 1021,697 size 32x24; Picture "Graphic_244"
   GraphicView "Graphic view_2" at 1021,558 size 32x24; Picture "Graphic_244"
   Button "HmiScreenItemData_1" at 1,1 size 150x43; TextOn 'Back'; TextOff 'Main Index'
      on Release: ActivateScreen("02 Main Index", 0)
   GraphicIOField "Graphic I/O field_3" at 586,670 size 60x65; PictureList "Pump Ani"
      ProcessValue <- "FW Pump Animation"
   Button "HmiScreenItemData_3" at 1129,1 size 150x43; TextOn 'I&A Compressor Ok'; TextOff 'Back'
      on Release: function_efd93a16()
   AlarmView "Alarm view_1" at 0,777 size 1280x23
   IOField "I/O field_21" at 617,211 size 90x25; FormatPattern 999999; Unit  h
      ProcessValue <- "P305_Functioning Hours_IDB_Hours Total"
      Visibility <- "80_From_HMI_P301_PRSNT"
   TextField "Text field_31" at 712,213 size 123x20; Text 'Total Run Hours'
      Visibility <- "80_From_HMI_P301_PRSNT"
   IOField "I/O field_1" at 648,173 size 40x25; FormatPattern 99; Unit d
      ProcessValue <- "82_To_HMI_P305 FW Pump Run Days"
   IOField "I/O field_9" at 646,273 size 65x25; Authorization "Commissioning"; FormatPattern 99999; Unit  h
      ProcessValue <- "82_To_HMI_P305 FW Pump Service Time Hours"
   Button "HmiScreenItemData_4" at 488,210 size 75x34; TextOn 'STOP'; TextOff 'Stop'
      on Press: ResetBit("80_From_HMI_MAN_DQ_1_7(1)")
   Button "HmiScreenItemData_2" at 385,210 size 75x34; TextOn 'START'; TextOff 'Start'
      on Press: SetBit("80_From_HMI_MAN_DQ_1_7(1)")
   Rectangle "Rectangle_7" at 208,78 size 656x250
      Visibility <- "80_From_HMI_P305_PRSNT"

screen "GCU Process Times" 1280x800, template "Template"
   on GenerateScreen: "TitleUpdater"()
   Button "HmiScreenItemData_1" at 1,1 size 150x43; TextOn 'Back'; TextOff 'Commissioning'
      on Release: ActivateScreen("Commissioning Main Page", 0)
   AlarmView "Alarm view_1" at 0,777 size 1280x23
   TextField "Text field_29" at 545,103 size 65x20; Text 'Time (s)'
   TextField "Text field_65" at 240,128 size 300x25; Text 'P303 Started Delay'
   TextField "Text field_42" at 240,103 size 89x20; Text 'Description'
   IOField "I/O field_128" at 545,128 size 65x25; Authorization "Parameter Change"; FormatPattern 999
      ProcessValue <- "86_Times_P303_STRTD_DLY"
   TextField "Text field_53" at 240,74 size 193x26; Text 'GCU Process Times'
   TextField "Text field_1" at 240,158 size 300x25; Text 'P303 Stopped Delay'
   IOField "I/O field_1" at 545,158 size 65x25; Authorization "Parameter Change"; FormatPattern 999
      ProcessValue <- "86_Times_P303_STPD_DLY"
   TextField "Text field_2" at 240,188 size 300x25; Text 'P304 Started Delay'
   IOField "I/O field_2" at 545,188 size 65x25; Authorization "Parameter Change"; FormatPattern 999
      ProcessValue <- "86_Times_P304_STRTD_DLY"
   TextField "Text field_3" at 240,218 size 300x25; Text 'P304 Stopped Delay'
   IOField "I/O field_3" at 545,218 size 65x25; Authorization "Parameter Change"; FormatPattern 999
      ProcessValue <- "86_Times_P304_STPD_DLY"
   TextField "Text field_4" at 240,248 size 300x25; Text 'P305 Started Delay'
   IOField "I/O field_4" at 545,248 size 65x25; Authorization "Parameter Change"; FormatPattern 999
      ProcessValue <- "86_Times_P305_STRTD_DLY"
   TextField "Text field_5" at 240,278 size 300x25; Text 'P305 Stopped Delay'
   IOField "I/O field_5" at 545,278 size 65x25; Authorization "Parameter Change"; FormatPattern 999
      ProcessValue <- "86_Times_P305_STPD_DLY"
   TextField "Text field_6" at 240,308 size 300x25; Text 'CV341 Closed Delay'
   IOField "I/O field_6" at 545,308 size 65x25; Authorization "Parameter Change"; FormatPattern 999
      ProcessValue <- "86_Times_CV341_CLSD_DLY"
   TextField "Text field_7" at 240,338 size 300x25; Text 'CV358 Closed Delay'
   IOField "I/O field_7" at 545,338 size 65x25; Authorization "Parameter Change"; FormatPattern 999
      ProcessValue <- "86_Times_CV358_CLSD_DLY"
   TextField "Text field_8" at 975,103 size 65x20; Text 'Time (s)'
   TextField "Text field_9" at 670,128 size 300x25; Text 'CV405 Opened Delay'
   TextField "Text field_10" at 670,103 size 89x20; Text 'Description'
   IOField "I/O field_8" at 975,128 size 65x25; Authorization "Parameter Change"; FormatPattern 999
      ProcessValue <- "86_Times_CV405_OPND_DLY"
   TextField "Text field_11" at 670,158 size 300x25; Text 'CV406 Closed Delay'
   IOField "I/O field_9" at 975,158 size 65x25; Authorization "Parameter Change"; FormatPattern 999
      ProcessValue <- "86_Times_CV406_CLSD_DLY"
   TextField "Text field_12" at 670,188 size 300x25; Text 'E400 Stop Time'
   IOField "I/O field_10" at 975,188 size 65x25; Authorization "Parameter Change"; FormatPattern 999
      ProcessValue <- "86_Times_E400_STOP_TIME"
   TextField "Text field_13" at 670,218 size 300x25; Text 'P303 Stop Time'
   IOField "I/O field_11" at 975,218 size 65x25; Authorization "Parameter Change"; FormatPattern 999
      ProcessValue <- "86_Times_P303_STOP_TIME"
   TextField "Text field_14" at 670,248 size 300x25; Text 'CV341 Opened Delay'
   IOField "I/O field_12" at 975,248 size 65x25; Authorization "Parameter Change"; FormatPattern 999
      ProcessValue <- "86_Times_CV341_OPND_DLY"
   TextField "Text field_15" at 670,278 size 300x25; Text 'GCU Tank Maximum Drain Time'
   IOField "I/O field_13" at 975,278 size 65x25; Authorization "Parameter Change"; FormatPattern 999
      ProcessValue <- "86_Times_GCU_TNK_DRN_MAX_TIME"
   TextField "Text field_16" at 670,308 size 300x25; Text 'GCU Flush Time'
   IOField "I/O field_14" at 975,308 size 65x25; Authorization "Parameter Change"; FormatPattern 999
      ProcessValue <- "86_Times_GCU_FLUSH_TIME"
   TextField "Text field_17" at 670,338 size 300x25; Text 'Post Flush Delay'
   IOField "I/O field_15" at 975,338 size 65x25; Authorization "Parameter Change"; FormatPattern 999
      ProcessValue <- "86_Times_POST_FLUSH_DLY"
   TextField "Text field_18" at 240,368 size 300x25; Text 'CV401 Opened Delay'
   IOField "I/O field_16" at 545,368 size 65x25; Authorization "Parameter Change"; FormatPattern 999
      ProcessValue <- "86_Times_CV401_OPND_DLY"
   TextField "Text field_19" at 240,398 size 300x25; Text 'CV401 Closed Delay'
   IOField "I/O field_17" at 545,398 size 65x25; Authorization "Parameter Change"; FormatPattern 999
      ProcessValue <- "86_Times_CV401_CLSD_DLY"
   TextField "Text field_20" at 240,428 size 300x25; Text 'CV441 Opened Delay'
   IOField "I/O field_18" at 545,428 size 65x25; Authorization "Parameter Change"; FormatPattern 999
      ProcessValue <- "86_Times_CV441_OPND_DLY"
   TextField "Text field_21" at 240,458 size 300x25; Text 'CV441 Closed Delay'
   IOField "I/O field_19" at 545,458 size 65x25; Authorization "Parameter Change"; FormatPattern 999
      ProcessValue <- "86_Times_CV441_CLSD_DLY"
   TextField "Text field_22" at 240,488 size 300x25; Text 'Pre CV441 Open Delay'
   IOField "I/O field_20" at 545,488 size 65x25; Authorization "Parameter Change"; FormatPattern 999
      ProcessValue <- "86_Times_PRE_CV441_OPN_DLY"
   TextField "Text field_23" at 240,518 size 300x25; Text 'Valve Configuration Done Delay'
   IOField "I/O field_21" at 545,518 size 65x25; Authorization "Parameter Change"; FormatPattern 999
      ProcessValue <- "86_Times_VLV_CNFG_DN_DLY"
   TextField "Text field_24" at 240,548 size 300x25; Text 'Pre GCU Tank Fill Delay'
   IOField "I/O field_22" at 545,548 size 65x25; Authorization "Parameter Change"; FormatPattern 999
      ProcessValue <- "86_Times_PRE_GCU_TNK_FILL_DLY"
   TextField "Text field_25" at 240,578 size 300x25; Text 'GCU Tank Fill Maximum Time'
   IOField "I/O field_23" at 545,578 size 65x25; Authorization "Parameter Change"; FormatPattern 999
      ProcessValue <- "86_Times_GCU_TNK_FILL_MAX_TIME"
   TextField "Text field_26" at 670,368 size 300x25; Text 'CV341 Maximum Travel Time'
   IOField "I/O field_24" at 975,368 size 65x25; Authorization "Parameter Change"; FormatPattern 999
      ProcessValue <- "86_Times_CV341_MAX_TRVL_TIME"
   TextField "Text field_27" at 670,398 size 300x25; Text 'CV358 Maximum Travel Time'
   IOField "I/O field_25" at 975,398 size 65x25; Authorization "Parameter Change"; FormatPattern 999
      ProcessValue <- "86_Times_CV358_MAX_TRVL_TIME"
   TextField "Text field_28" at 670,428 size 300x25; Text 'CV406 Maximum Travel Time'
   IOField "I/O field_26" at 975,428 size 65x25; Authorization "Parameter Change"; FormatPattern 999
      ProcessValue <- "86_Times_CV406_MAX_TRVL_TIME"
   TextField "Text field_30" at 670,458 size 300x25; Text 'CV407 Maximum Travel Time'
   IOField "I/O field_27" at 975,458 size 65x25; Authorization "Parameter Change"; FormatPattern 999
      ProcessValue <- "86_Times_CV407_MAX_TRVL_TIME"
   TextField "Text field_31" at 670,488 size 300x25; Text 'CV409 Maximum Travel Time'
   IOField "I/O field_28" at 975,488 size 65x25; Authorization "Parameter Change"; FormatPattern 999
      ProcessValue <- "86_Times_CV409_MAX_TRVL_TIME"
   TextField "Text field_32" at 670,518 size 300x25; Text 'CV411 Maximum Travel Time'
   IOField "I/O field_29" at 975,518 size 65x25; Authorization "Parameter Change"; FormatPattern 999
      ProcessValue <- "86_Times_CV411_MAX_TRVL_TIME"
   TextField "Text field_33" at 670,548 size 300x25; Text 'CV441 Maximum Travel Time'
   IOField "I/O field_30" at 975,548 size 65x25; Authorization "Parameter Change"; FormatPattern 999
      ProcessValue <- "86_Times_CV441_MAX_TRVL_TIME"
   TextField "Text field_34" at 670,638 size 300x25; Text 'PIT416 Target Ramp Time'
   IOField "I/O field_31" at 975,638 size 65x25; Authorization "Parameter Change"; FormatPattern 999
      ProcessValue <- "86_Times_PIT416_TRGT_RMP_TIME"
   TextField "Text field_35" at 240,608 size 300x25; Text 'E400 Started Delay'
   IOField "I/O field_32" at 545,608 size 65x25; Authorization "Parameter Change"; FormatPattern 999
      ProcessValue <- "86_Times_E400_STRTD_DLY"
   TextField "Text field_36" at 240,638 size 300x25; Text 'E400 Running Delay'
   IOField "I/O field_33" at 545,638 size 65x25; Authorization "Parameter Change"; FormatPattern 999
      ProcessValue <- "86_Times_E400_RNG_DLY"
   TextField "Text field_37" at 670,578 size 300x25; Text 'PIT353 Alarm Delay Time'
   IOField "I/O field_34" at 975,578 size 65x25; Authorization "Parameter Change"; FormatPattern 999
      ProcessValue <- "86_Times_PIT353 Delay"
   TextField "Text field_38" at 670,608 size 300x25; Text 'PIT416 Alarm Delay Time'
   IOField "I/O field_35" at 975,608 size 65x25; Authorization "Parameter Change"; FormatPattern 999
      ProcessValue <- "86_Times_PIT416 Delay"
   TextField "Text field_39" at 240,669 size 300x25; Text 'P301 Started Delay'
   IOField "I/O field_36" at 545,669 size 65x25; Authorization "Parameter Change"; FormatPattern 999
      ProcessValue <- "86_Times_P301_START_DLY"
   TextField "Text field_40" at 670,669 size 300x25; Text 'FS332 Alarm Delay'
   IOField "I/O field_37" at 975,669 size 65x25; Authorization "Parameter Change"; FormatPattern 999
      ProcessValue <- "86_Times_FS332 Delay"
   TextField "Text field_41" at 670,701 size 300x25; Text 'LIT304 Alarm Delay'
   IOField "I/O field_38" at 975,701 size 65x25; Authorization "Parameter Change"; FormatPattern 999
      ProcessValue <- "86_Times_LIT304 Delay"
   Group "Group" at 455,41 size 373x50
   TextField "Text field_43" at 240,701 size 300x25; Text 'PIT358 Alarm Delay Time'
   IOField "I/O field_39" at 545,701 size 65x25; Authorization "Parameter Change"; FormatPattern 999
      ProcessValue <- "86_Times_PIT358 Delay"
   TextField "Text field_44" at 240,732 size 300x25; Text 'PIT348 Alarm Delay Time'
   IOField "I/O field_40" at 545,732 size 65x25; Authorization "Parameter Change"; FormatPattern 999
      ProcessValue <- "86_Times_PIT348 Delay"
   Button "HmiScreenItemData_8" at 469,45 size 355x40; TextOn 'Back'; TextOff 'Text'
   TextField "Screen title" at 455,41 size 373x50; Text 'Screen title'

Template "Template_lite" 1280x800
   Button "HmiScreenItemData_12" at 993,4 size 80x35; TextOn 'WARNING'; TextOff 'Warning'
      on Release: ActivateScreen("04 Alarm Log", 0)
      Visibility <- "62_Warning_Data_WRNG_PRSNT"
   Button "HmiScreenItemData_14" at 1080,4 size 80x35; TextOn 'ALARM'; TextOff 'Alarm'
      on Release: ActivateScreen("04 Alarm Log", 0)
      Visibility <- "60_Alarm_Data_ALRM_PRSNT"
   Button "HmiScreenItemData_20" at 906,4 size 80x35; TextOn 'Back'; TextOff 'Lockout'
      on Click: SetBit("80_From_HMI_Reset_Alarms")
      on Press: function_b14e0dd5("80_From_HMI_RST_LOCKOUT", 0)
      Appearance <- "82_To_HMI_E-STOP LATCHED"
   Button "HmiScreenItemData_24" at 810,3 size 64x35; TextOn 'MUTE'; TextOff 'Mute'
      on Press: function_b14e0dd5("80_From_HMI_SLNCE_BZR", 0)
      Appearance <- "80_From_HMI_SLNCE_BZR"
   GraphicView "Graphic view_24" at 876,3 size 29x41; Picture "Graphic_138"
      Visibility <- "Buzzer"
   Circle "Circle_46" at 265,6 size 26x26
      Visibility <- "TRUE"
      Appearance <- "IGG PLC HEART BEAT"
   Circle "Circle_1" at 235,6 size 26x26
      Visibility <- "TRUE"
      Appearance <- "Setpoint Override_DB_Set Pressure"

